// TIA Portal project "SemesterprosjektV7" (V20)

(* hardware
DEVICE "S7-1200 station_1"  S7-1200 Station
   slot 0: "Rack_0"  S7-1200 Rack  Rack  V1.0
   slot 1: "PLC_1"  CPU 1212C AC/DC/Rly  6ES7 212-1BD30-0XB0  V2.0
   slot 2: "AI 4x13BIT_1"  SM 1231 AI4  6ES7 231-4HD32-0XB0  V2.1
   slot 3: "AQ 2x14BIT_1"  SM 1232 AQ2  6ES7 232-4HB32-0XB0  V2.1
DEVICE "HMI_1"  KTP700 Basic PN
   slot 0: "HMI_1"  KTP700 Basic PN  6AV2 123-2GB03-0AX0  17.0.0.0
   slot 1: "HMI_RT_1"  KTP700 Basic PN  6AV2 123-2GB03-0AX0  17.0.0.0
   slot 5: "HMI_1.IE_CP_1"  PROFINET Interface  17.0.0.0
      slot 1: "PROFINET Interface_1"  PROFINET Interface
         slot 1: "Port_1"  Port
*)

// ===== PLC "PLC_1"  CPU 1212C AC/DC/Rly =====

VAR_GLOBAL   // PLC tag table "Default tag table"
   "AI2+" AT %IW100 : Int;
   "AQ1_PÅDRAG_PUMP1" AT %QW112 : Int;
   "AQ2" AT %QW114 : Int;
   "DI_EM_STOP" AT %I0.0 : Bool;
   "DQ_START_PUMP1" AT %Q0.0 : Bool;
   "DI_LS_Tørrkjøringsvern" AT %I0.1 : Bool;
   "DI_Reset_EM_STOP" AT %I0.2 : Bool;
   "DQ_Lys_EM_STOP" AT %Q0.1 : Bool;
END_VAR

// folder: Equipment

TYPE "UDT_Mal"
   STRUCT
      CFG : Struct   // Configuration Data
         Spare : Bool;
      END_STRUCT;
      Sts : Struct   // Status Data
         Spare : Bool;
      END_STRUCT;
      Cmd : Struct   // Command and request Data
         Spare : Bool;
      END_STRUCT;
      Par : Struct   // Parameter Data
         Spare : Bool;
      END_STRUCT;
      Fit : Struct   // Warning and alarm triggers
         Spare : Bool;
      END_STRUCT;
   END_STRUCT;
END_TYPE

TYPE "UDT_Pump_Control"
   STRUCT
      CFG : Struct   // Configuration Data
         Spare : Bool;
      END_STRUCT;
      Sts : Struct   // Status Data
         Spare : Bool;
      END_STRUCT;
      Cmd : Struct   // Command and request Data
         Start_Pump : Bool;
         Stop_Pump : Bool;
         EM_Stop : Bool;
      END_STRUCT;
      Par : Struct   // Parameter Data
         Pådrag_Inn : Real;
      END_STRUCT;
      Fit : Struct   // Warning and alarm triggers
         Feil : Bool;
      END_STRUCT;
   END_STRUCT;
END_TYPE

TYPE "UDT_Level_Transmitter"
   STRUCT
      CFG : Struct   // Configuration Data
         Spare : Bool;
      END_STRUCT;
      Sts : Struct   // Status Data
         Spare : Bool;
      END_STRUCT;
      Cmd : Struct   // Command and request Data
         Spare : Bool;
      END_STRUCT;
      Par : Struct   // Parameter Data
         EU_Value_Out : Real;
      END_STRUCT;
      Fit : Struct   // Warning and alarm triggers
         Feil : Bool;
         Spare : Bool;
      END_STRUCT;
   END_STRUCT;
END_TYPE

// folder: Machine

TYPE "UDT_HMI"
   STRUCT
      CFG : Struct   // Configuration Data
         Spare : Bool;
      END_STRUCT;
      Sts : Struct   // Status Data
         HMI_Level_PV : Real;
      END_STRUCT;
      Cmd : Struct   // Command and request Data
         HMI_Auto : Bool;
         HMI_Manuell : Bool;
         HMI_Start_Pump1 : Bool;
         HMI_Stop_Pump1 : Bool;
         HMI_Knapp_Auto : Bool;
         HMI_Knapp_Manuell : Bool;
         HMI_Knapp_Start_Pump1 : Bool;
         HMI_Knapp_Stop_Pump1 : Bool;
         Spare : Bool;
      END_STRUCT;
      Par : Struct   // Parameter Data
         HMI_P_Gain : Real;
         HMI_Ti : Real;
         HMI_Td : Real;
         HMI_Manual_Speed_Ref_P1 : Real;
         HMI_Level_SP : Real;
         HMI_EU_Min : Real;
         HMI_EU_Max : Real;
         HMI_Anti_Windup : Bool;
         Spare : Bool;
      END_STRUCT;
      Fit : Struct   // Warning and alarm triggers
         HMI_EM_Stop_Alarm : Bool;
         HMI_LS_Activated : Bool;
         HMI_Pump_Fault_Timer_SP : Time;
         HMI_Pump_Fault : Bool;
         Spare : Bool;
      END_STRUCT;
   END_STRUCT;
END_TYPE

// folder: (top level)

DATA_BLOCK "LT01"   // DB3
{ S7_Optimized_Access := 'TRUE' }
VERSION : 0.1
// stored: InstanceOfName Level_Transmitter
"Level_Transmitter"
BEGIN
END_DATA_BLOCK

DATA_BLOCK "Analog_Data"   // DB4
{ S7_Optimized_Access := 'TRUE' }
VERSION : 0.1
   VAR
      Raw_Value : Real;
      Output : Real;
      EU_Min : Real;
      EU_Max : Real;
   END_VAR
BEGIN
END_DATA_BLOCK

DATA_BLOCK "Pump1_Control_DB"   // DB6
{ S7_Optimized_Access := 'TRUE' }
VERSION : 0.1
// stored: InstanceOfName Pump_Control
"Pump_Control"
BEGIN
END_DATA_BLOCK

DATA_BLOCK "Machine01_DB"   // DB7
{ S7_Optimized_Access := 'TRUE' }
VERSION : 0.1
// stored: InstanceOfName Machine01
"Machine01"
BEGIN
END_DATA_BLOCK

DATA_BLOCK "Regulator_DB"   // DB9
{ S7_Optimized_Access := 'TRUE' }
VERSION : 0.1
// stored: InstanceOfName Regulator
"Regulator"
BEGIN
END_DATA_BLOCK

// folder: Global_Data

DATA_BLOCK "DB_Machine"   // DB1
{ S7_Optimized_Access := 'TRUE' }
VERSION : 0.1
   VAR
      HMI_Control : "UDT_HMI";
   END_VAR
BEGIN
END_DATA_BLOCK

DATA_BLOCK "DB_Equipment"   // DB2
{ S7_Optimized_Access := 'TRUE' }
VERSION : 0.1
   VAR
      Pump1_Control : "UDT_Pump_Control";
      LT01_Control : "UDT_Level_Transmitter";
      HMI_Control : "UDT_HMI";
   END_VAR
BEGIN
END_DATA_BLOCK

// folder: System blocks/Program resources

DATA_BLOCK "EM_Stop_TON_DB"   // DB5
{ S7_Optimized_Access := 'TRUE' }
AUTHOR : Simatic
FAMILY : IEC
NAME : IEC_TMR
VERSION : 1.0
// stored: InstanceOfName IEC_TIMER
"IEC_TIMER"
BEGIN
END_DATA_BLOCK

DATA_BLOCK "EM_Stop_TOF_DB"   // DB10
{ S7_Optimized_Access := 'TRUE' }
AUTHOR : Simatic
FAMILY : IEC
NAME : IEC_TMR
VERSION : 1.0
// stored: InstanceOfName IEC_TIMER
"IEC_TIMER"
BEGIN
END_DATA_BLOCK

DATA_BLOCK "Pump_Fault_Timer_DB"   // DB11
{ S7_Optimized_Access := 'TRUE' }
AUTHOR : Simatic
FAMILY : IEC
NAME : IEC_TMR
VERSION : 1.0
// stored: InstanceOfName IEC_TIMER
"IEC_TIMER"
BEGIN
END_DATA_BLOCK

// folder: (top level)

ORGANIZATION_BLOCK "Main"   // OB1, LAD, ProgramCycle
TITLE = "Main Program Sweep (Cycle)"
{ S7_Optimized_Access := 'TRUE' }
VERSION : 0.1
BEGIN
END_ORGANIZATION_BLOCK

ORGANIZATION_BLOCK "Machine"   // OB123, LAD, ProgramCycle
TITLE = "Main Program Sweep (Cycle)"
{ S7_Optimized_Access := 'TRUE' }
VERSION : 0.1
BEGIN

REGION Network 1
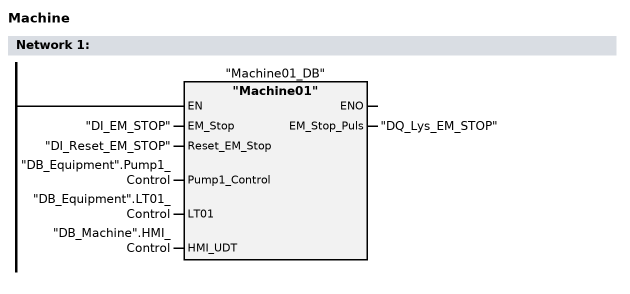
   RUNG wire#powerrail
      "Machine01_DB"(EM_Stop := "DI_EM_STOP", Reset_EM_Stop := "DI_Reset_EM_STOP", Pump1_Control := "DB_Equipment".Pump1_Control, LT01 := "DB_Equipment".LT01_Control, HMI_UDT := "DB_Machine".HMI_Control, EM_Stop_Puls => "DQ_Lys_EM_STOP")
   END_RUNG
   // the same network as SCL:
   "Machine01_DB"(EM_Stop := "DI_EM_STOP",   // "Machine01"
                  Reset_EM_Stop := "DI_Reset_EM_STOP",
                  Pump1_Control := "DB_Equipment".Pump1_Control,
                  LT01 := "DB_Equipment".LT01_Control,
                  HMI_UDT := "DB_Machine".HMI_Control,
                  EM_Stop_Puls => "DQ_Lys_EM_STOP");
END_REGION
END_ORGANIZATION_BLOCK

ORGANIZATION_BLOCK "Equipment"   // OB124, LAD, ProgramCycle
TITLE = "Main Program Sweep (Cycle)"
{ S7_Optimized_Access := 'TRUE' }
VERSION : 0.1
BEGIN

REGION Network 1
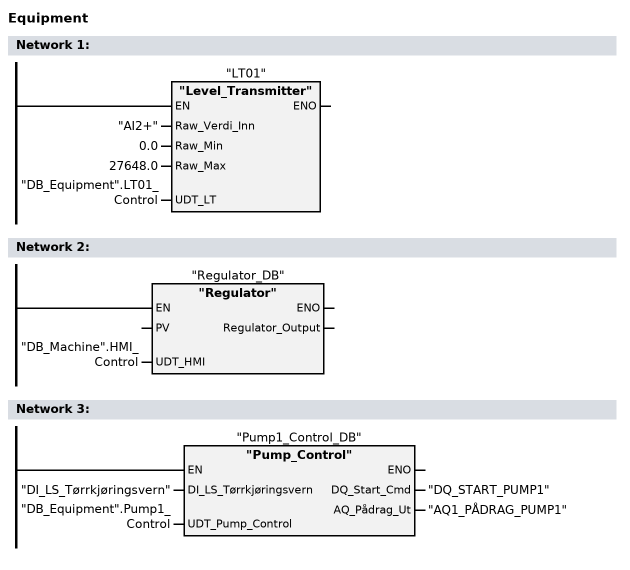
   RUNG wire#powerrail
      "LT01"(Raw_Verdi_Inn := "AI2+", Raw_Min := 0.0, Raw_Max := 27648.0, UDT_LT := "DB_Equipment".LT01_Control)
   END_RUNG
   // the same network as SCL:
   "LT01"(Raw_Verdi_Inn := "AI2+", Raw_Min := 0.0, Raw_Max := 27648.0, UDT_LT := "DB_Equipment".LT01_Control);   // "Level_Transmitter"
END_REGION

REGION Network 2
   RUNG wire#powerrail
      "Regulator_DB"(PV :=, UDT_HMI := "DB_Machine".HMI_Control, Regulator_Output =>)
   END_RUNG
   // the same network as SCL:
   "Regulator_DB"(UDT_HMI := "DB_Machine".HMI_Control);   // "Regulator"
END_REGION

REGION Network 3
   RUNG wire#powerrail
      "Pump1_Control_DB"(DI_LS_Tørrkjøringsvern := "DI_LS_Tørrkjøringsvern", UDT_Pump_Control := "DB_Equipment".Pump1_Control, DQ_Start_Cmd => "DQ_START_PUMP1", AQ_Pådrag_Ut => "AQ1_PÅDRAG_PUMP1")
   END_RUNG
   // the same network as SCL:
   "Pump1_Control_DB"(DI_LS_Tørrkjøringsvern := "DI_LS_Tørrkjøringsvern",   // "Pump_Control"
                      UDT_Pump_Control := "DB_Equipment".Pump1_Control,
                      DQ_Start_Cmd => "DQ_START_PUMP1",
                      AQ_Pådrag_Ut => "AQ1_PÅDRAG_PUMP1");
END_REGION
END_ORGANIZATION_BLOCK

// folder: Equipment

FUNCTION_BLOCK "Pump_Control"   // FB2, LAD
{ S7_Optimized_Access := 'TRUE' }
VERSION : 0.1
   VAR_INPUT
      DI_LS_Tørrkjøringsvern : Bool;
   END_VAR
   VAR_OUTPUT
      DQ_Start_Cmd : Bool;
      AQ_Pådrag_Ut : Int;
   END_VAR
   VAR_IN_OUT
      UDT_Pump_Control : "UDT_Pump_Control";
   END_VAR
   VAR
      Tmp_Start_Cmd : Bool;
      Tmp_Pådrag_Ut_Real : Real;
      Temp_Verdi : Real;
      Tmp_Pådrag_Ut_Int : Real;
   END_VAR
BEGIN

REGION Network 1
   // Start Pumpe og stopp kriterier
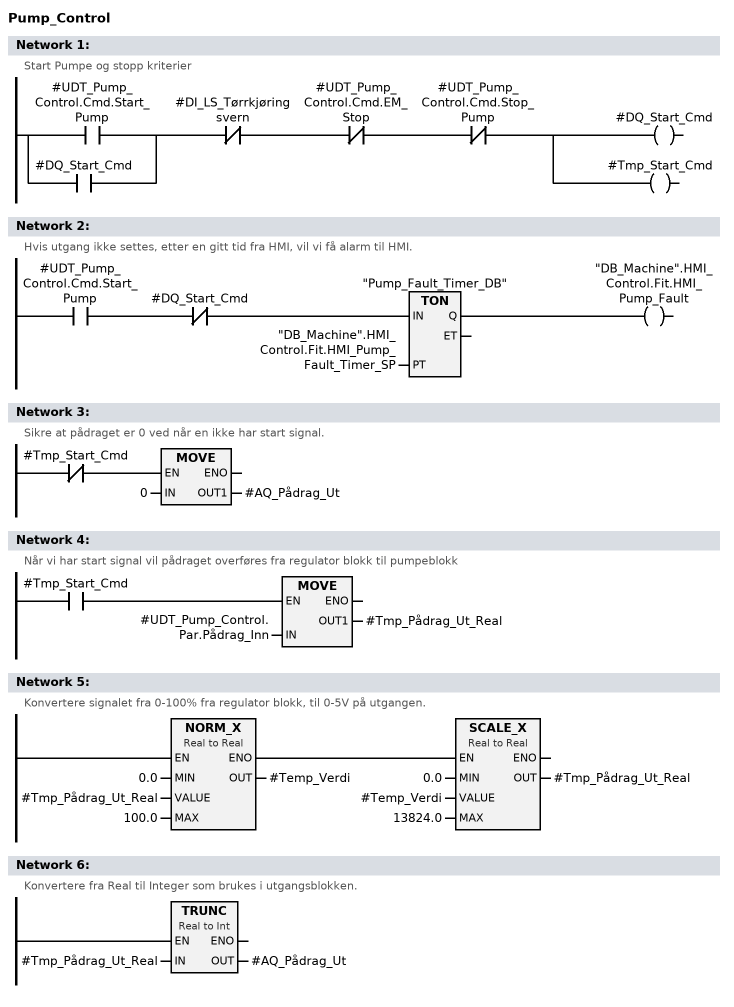
   RUNG wire#powerrail
      Contact( #UDT_Pump_Control.Cmd.Start_Pump )
      wire#w1
      I_Contact( #DI_LS_Tørrkjøringsvern )
      I_Contact( #UDT_Pump_Control.Cmd.EM_Stop )
      I_Contact( #UDT_Pump_Control.Cmd.Stop_Pump )
      wire#w2
      Coil( #DQ_Start_Cmd )
   END_RUNG
   RUNG wire#powerrail
      Contact( #DQ_Start_Cmd )
   END_RUNG wire#w1
   RUNG wire#w2
      Coil( #Tmp_Start_Cmd )
   END_RUNG
   // the same network as SCL:
   #DQ_Start_Cmd := (#UDT_Pump_Control.Cmd.Start_Pump OR #DQ_Start_Cmd) AND NOT #DI_LS_Tørrkjøringsvern AND NOT #UDT_Pump_Control.Cmd.EM_Stop AND NOT #UDT_Pump_Control.Cmd.Stop_Pump;
   #Tmp_Start_Cmd := #DQ_Start_Cmd;
END_REGION

REGION Network 2
   // Hvis utgang ikke settes, etter en gitt tid fra HMI, vil vi få alarm til HMI.
   "Pump_Fault_Timer_DB".TON(IN := #UDT_Pump_Control.Cmd.Start_Pump AND NOT #DQ_Start_Cmd,
                           PT := "DB_Machine".HMI_Control.Fit.HMI_Pump_Fault_Timer_SP);
   "DB_Machine".HMI_Control.Fit.HMI_Pump_Fault := "Pump_Fault_Timer_DB".Q;
END_REGION

REGION Network 3
   // Sikre at pådraget er 0 ved når en ikke har start signal.
   RUNG wire#powerrail
      I_Contact( #Tmp_Start_Cmd )
      { S7_GenerateENO := "TRUE" } Move(in := 0, out1 => #AQ_Pådrag_Ut)
   END_RUNG
   // the same network as SCL:
   IF NOT #Tmp_Start_Cmd THEN #AQ_Pådrag_Ut := 0; END_IF;
END_REGION

REGION Network 4
   // Når vi har start signal vil pådraget overføres fra regulator blokk til pumpeblokk
   RUNG wire#powerrail
      Contact( #Tmp_Start_Cmd )
      { S7_GenerateENO := "TRUE" } Move(in := #UDT_Pump_Control.Par.Pådrag_Inn, out1 => #Tmp_Pådrag_Ut_Real)
   END_RUNG
   // the same network as SCL:
   IF #Tmp_Start_Cmd THEN #Tmp_Pådrag_Ut_Real := #UDT_Pump_Control.Par.Pådrag_Inn; END_IF;
END_REGION

REGION Network 5
   // Konvertere signalet fra 0-100% fra regulator blokk, til 0-5V på utgangen.
   RUNG wire#powerrail
      { S7_Templates := "[SrcType := Real, DestType := Real]"; S7_GenerateENO := "TRUE" } Normalize(min := 0.0, value := #Tmp_Pådrag_Ut_Real, max := 100.0, out => #Temp_Verdi)
      { S7_Templates := "[SrcType := Real, DestType := Real]"; S7_GenerateENO := "TRUE" } Scale(min := 0.0, value := #Temp_Verdi, max := 13824.0, out => #Tmp_Pådrag_Ut_Real)
   END_RUNG
   // the same network as SCL:
   // ENO of a box is taken as its EN; it also drops when the box reports an error
   #Temp_Verdi := NORM_X(MIN := 0.0, VALUE := #Tmp_Pådrag_Ut_Real, MAX := 100.0);
   #Tmp_Pådrag_Ut_Real := SCALE_X(MIN := 0.0, VALUE := #Temp_Verdi, MAX := 13824.0);
END_REGION

REGION Network 6
   // Konvertere fra Real til Integer som brukes i utgangsblokken.
   RUNG wire#powerrail
      { S7_Templates := "[SrcType := Real, DestType := Int]"; S7_GenerateENO := "TRUE" } Trunc(in := #Tmp_Pådrag_Ut_Real, out => #AQ_Pådrag_Ut)
   END_RUNG
   // the same network as SCL:
   #AQ_Pådrag_Ut := TRUNC(#Tmp_Pådrag_Ut_Real);
END_REGION
END_FUNCTION_BLOCK

FUNCTION_BLOCK "Level_Transmitter"   // FB3, LAD
{ S7_Optimized_Access := 'TRUE' }
VERSION : 0.1
   VAR_INPUT
      Raw_Verdi_Inn : Int;
      Raw_Min : Real;
      Raw_Max : Real;
   END_VAR
   VAR_IN_OUT
      UDT_LT : "UDT_Level_Transmitter";
   END_VAR
   VAR_TEMP
      Convert_Value : Real;
      Raw_Value_Real : Real;
   END_VAR
BEGIN

REGION Network 1
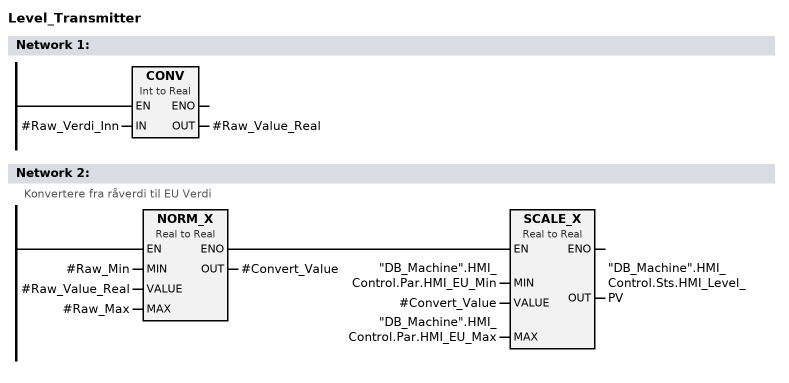
   RUNG wire#powerrail
      { S7_Templates := "[SrcType := Int, DestType := Real]"; S7_GenerateENO := "TRUE" } Convert(in := #Raw_Verdi_Inn, out => #Raw_Value_Real)
   END_RUNG
   // the same network as SCL:
   #Raw_Value_Real := INT_TO_REAL(#Raw_Verdi_Inn);
END_REGION

REGION Network 2
   // Konvertere fra råverdi til EU Verdi
   RUNG wire#powerrail
      { S7_Templates := "[SrcType := Real, DestType := Real]"; S7_GenerateENO := "TRUE" } Normalize(min := #Raw_Min, value := #Raw_Value_Real, max := #Raw_Max, out => #Convert_Value)
      { S7_Templates := "[SrcType := Real, DestType := Real]"; S7_GenerateENO := "TRUE" } Scale(min := "DB_Machine".HMI_Control.Par.HMI_EU_Min, value := #Convert_Value, max := "DB_Machine".HMI_Control.Par.HMI_EU_Max, out => "DB_Machine".HMI_Control.Sts.HMI_Level_PV)
   END_RUNG
   // the same network as SCL:
   // ENO of a box is taken as its EN; it also drops when the box reports an error
   #Convert_Value := NORM_X(MIN := #Raw_Min, VALUE := #Raw_Value_Real, MAX := #Raw_Max);
   "DB_Machine".HMI_Control.Sts.HMI_Level_PV := SCALE_X(MIN := "DB_Machine".HMI_Control.Par.HMI_EU_Min, VALUE := #Convert_Value, MAX := "DB_Machine".HMI_Control.Par.HMI_EU_Max);
END_REGION
END_FUNCTION_BLOCK

FUNCTION_BLOCK "ØL_PID"   // FB4, LAD
{ S7_Optimized_Access := 'TRUE' }
VERSION : 0.1
   VAR_INPUT
      SP : LReal;   // // NRM / SIU Setpoint
      PV : LReal;   // // NRM / SIU Process Value
      Bias : LReal;   // // NRM Bias Value
      I_SP : LReal;   // // NRM Setpoint for integrator value
      I_SP_Cmd : Bool;   // // TRUE: Load I_SP
      Suspend : Bool;   // // TRUE: Suspends operation
   END_VAR
   VAR_OUTPUT
      EV : LReal;   // // NRM / SIU Error Value
      CV : LReal;   // // NRM Control Value
   END_VAR
BEGIN
END_FUNCTION_BLOCK

FUNCTION_BLOCK "Regulator"   // FB5, LAD
{ S7_Optimized_Access := 'TRUE' }
VERSION : 0.1
   VAR_INPUT
      PV : Real;
   END_VAR
   VAR_OUTPUT
      Regulator_Output : Real;
   END_VAR
   VAR_IN_OUT
      UDT_HMI : "UDT_HMI";
   END_VAR
   VAR
      Convert_Value : Real;
      "Regulator_PV_%" : Real;
   END_VAR
BEGIN

REGION Network 2
   // Konvertere fra råverdi til EU Verdi
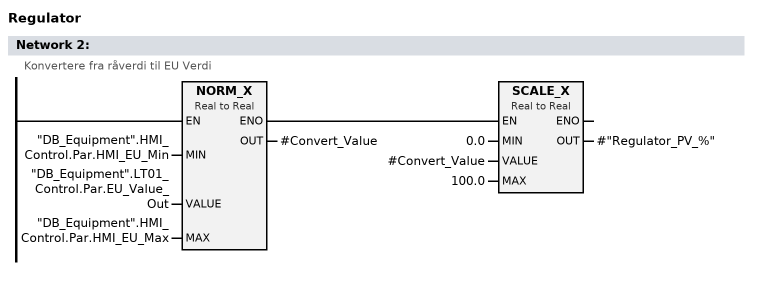
   RUNG wire#powerrail
      { S7_Templates := "[SrcType := Real, DestType := Real]"; S7_GenerateENO := "TRUE" } Normalize(min := "DB_Equipment".HMI_Control.Par.HMI_EU_Min, value := "DB_Equipment".LT01_Control.Par.EU_Value_Out, max := "DB_Equipment".HMI_Control.Par.HMI_EU_Max, out => #Convert_Value)
      { S7_Templates := "[SrcType := Real, DestType := Real]"; S7_GenerateENO := "TRUE" } Scale(min := 0.0, value := #Convert_Value, max := 100.0, out => #"Regulator_PV_%")
   END_RUNG
   // the same network as SCL:
   // ENO of a box is taken as its EN; it also drops when the box reports an error
   #Convert_Value := NORM_X(MIN := "DB_Equipment".HMI_Control.Par.HMI_EU_Min, VALUE := "DB_Equipment".LT01_Control.Par.EU_Value_Out, MAX := "DB_Equipment".HMI_Control.Par.HMI_EU_Max);
   #"Regulator_PV_%" := SCALE_X(MIN := 0.0, VALUE := #Convert_Value, MAX := 100.0);
END_REGION
END_FUNCTION_BLOCK

// folder: Machine

FUNCTION_BLOCK "Machine01"   // FB1, LAD
{ S7_Optimized_Access := 'TRUE' }
VERSION : 0.1
   VAR_INPUT
      EM_Stop : Bool;
      Reset_EM_Stop : Bool;
   END_VAR
   VAR_OUTPUT
      EM_Stop_Puls : Bool;
   END_VAR
   VAR_IN_OUT
      Pump1_Control : "UDT_Pump_Control";
      LT01 : "UDT_Level_Transmitter";
      HMI_UDT : "UDT_HMI";
   END_VAR
   VAR
      Tmp_EM_Stop : Bool;
      Tmp_Enable_PID : Bool;
      Tmp_Blink_Off : Bool;
      Tmp_Blink_On : Bool;
   END_VAR
BEGIN

REGION Network 1
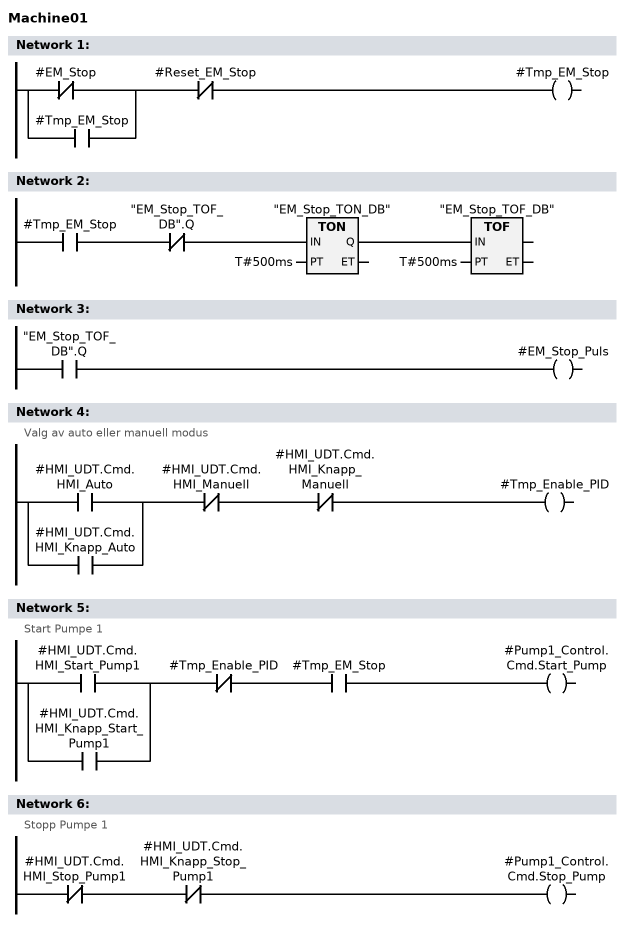
   RUNG wire#powerrail
      I_Contact( #EM_Stop )
      wire#w1
      I_Contact( #Reset_EM_Stop )
      Coil( #Tmp_EM_Stop )
   END_RUNG
   RUNG wire#powerrail
      Contact( #Tmp_EM_Stop )
   END_RUNG wire#w1
   // the same network as SCL:
   #Tmp_EM_Stop := (NOT #EM_Stop OR #Tmp_EM_Stop) AND NOT #Reset_EM_Stop;
END_REGION

REGION Network 2
   "EM_Stop_TON_DB".TON(IN := #Tmp_EM_Stop AND NOT "EM_Stop_TOF_DB".Q, PT := T#500ms);
   "EM_Stop_TOF_DB".TOF(IN := "EM_Stop_TON_DB".Q, PT := T#500ms);
END_REGION

REGION Network 3
   RUNG wire#powerrail
      Contact( "EM_Stop_TOF_DB".Q )
      Coil( #EM_Stop_Puls )
   END_RUNG
   // the same network as SCL:
   #EM_Stop_Puls := "EM_Stop_TOF_DB".Q;
END_REGION

REGION Network 4
   // Valg av auto eller manuell modus
   RUNG wire#powerrail
      Contact( #HMI_UDT.Cmd.HMI_Auto )
      wire#w1
      I_Contact( #HMI_UDT.Cmd.HMI_Manuell )
      I_Contact( #HMI_UDT.Cmd.HMI_Knapp_Manuell )
      Coil( #Tmp_Enable_PID )
   END_RUNG
   RUNG wire#powerrail
      Contact( #HMI_UDT.Cmd.HMI_Knapp_Auto )
   END_RUNG wire#w1
   // the same network as SCL:
   #Tmp_Enable_PID := (#HMI_UDT.Cmd.HMI_Auto OR #HMI_UDT.Cmd.HMI_Knapp_Auto) AND NOT #HMI_UDT.Cmd.HMI_Manuell AND NOT #HMI_UDT.Cmd.HMI_Knapp_Manuell;
END_REGION

REGION Network 5
   // Start Pumpe 1
   RUNG wire#powerrail
      Contact( #HMI_UDT.Cmd.HMI_Start_Pump1 )
      wire#w1
      I_Contact( #Tmp_Enable_PID )
      Contact( #Tmp_EM_Stop )
      Coil( #Pump1_Control.Cmd.Start_Pump )
   END_RUNG
   RUNG wire#powerrail
      Contact( #HMI_UDT.Cmd.HMI_Knapp_Start_Pump1 )
   END_RUNG wire#w1
   // the same network as SCL:
   #Pump1_Control.Cmd.Start_Pump := (#HMI_UDT.Cmd.HMI_Start_Pump1 OR #HMI_UDT.Cmd.HMI_Knapp_Start_Pump1) AND NOT #Tmp_Enable_PID AND #Tmp_EM_Stop;
END_REGION

REGION Network 6
   // Stopp Pumpe 1
   RUNG wire#powerrail
      I_Contact( #HMI_UDT.Cmd.HMI_Stop_Pump1 )
      I_Contact( #HMI_UDT.Cmd.HMI_Knapp_Stop_Pump1 )
      Coil( #Pump1_Control.Cmd.Stop_Pump )
   END_RUNG
   // the same network as SCL:
   #Pump1_Control.Cmd.Stop_Pump := NOT #HMI_UDT.Cmd.HMI_Stop_Pump1 AND NOT #HMI_UDT.Cmd.HMI_Knapp_Stop_Pump1;
END_REGION
END_FUNCTION_BLOCK

(* ===== HMI "HMI_RT_1" =====
system functions are stored by id; their names below are inferred from use
connection "HMI_Connection_1": ETHERNET, SMART_S7_1200_OMS

HMI tags "HMI_Tags"
   "Knapp_HMI_Stop_Pump1" : Bool = PLC DB_Machine.HMI_Control.Cmd.HMI_Knapp_Stop_Pump1 AT %DB1.DBX0.0, 1 s
   "HMI_Manuell" : Bool = PLC DB_Machine.HMI_Control.Cmd.HMI_Manuell AT %DB1.DBX0.0, 1 s
   "HMI_Start_Pump1" : Bool = PLC DB_Machine.HMI_Control.Cmd.HMI_Start_Pump1 AT %DB1.DBX0.0, 1 s
   "Knapp_HMI_Auto" : Bool = PLC DB_Machine.HMI_Control.Cmd.HMI_Knapp_Auto AT %DB1.DBX0.0, 1 s
   "HMI_Auto" : Bool = PLC DB_Machine.HMI_Control.Cmd.HMI_Auto AT %DB1.DBX0.0, 1 s
   "Knapp_HMI_Manuell" : Bool = PLC DB_Machine.HMI_Control.Cmd.HMI_Knapp_Manuell AT %DB1.DBX0.0, 1 s
   "Knapp_HMI_Start_Pump1" : Bool = PLC DB_Machine.HMI_Control.Cmd.HMI_Knapp_Start_Pump1 AT %DB1.DBX0.0, 1 s
   "Tag_ScreenNumber_1" : UInt, internal
   "HMI_Stop_Pump1" : Bool = PLC DB_Machine.HMI_Control.Cmd.HMI_Stop_Pump1 AT %DB1.DBX0.0, 1 s
   "PID_Compact_1_Output" : Real = PLC PID_Compact_1.Output, 1 s
   "PID_Compact_1_Setpoint" : Real = PLC PID_Compact_1.Setpoint, 1 s

Template "Template_1" 800x480
   Button "Exit" at 714,429 size 71x50; TextOff 'Exit'; PictureOff "ExitRuntime_KTP700_Basic_PN_TR"; PictureOn "ExitRuntime_KTP700_Basic_PN_TR"
      on Release: StopRuntime(0)
   Button "Log on" at 614,429 size 71x50; TextOff 'Log on'; PictureOff "Login_KTP700_Basic_PN_TR"; PictureOn "Login_KTP700_Basic_PN_TR"
      on Release: function_a2a04561()
   Button "Template_Button" at 514,429 size 71x50; TextOff 'Text'
   Button "Template_Button_1" at 414,429 size 71x50; TextOff 'Text'
   Button "Template_Button_2" at 314,429 size 71x50; TextOff 'Text'
   Button "Template_Button_3" at 214,429 size 71x50; TextOff 'Text'
   Button "Alarms" at 114,429 size 71x50; TextOff 'Alarms'; PictureOff "AlarmDisplay_KTP700_Basic_PN_TR"; PictureOn "AlarmDisplay_KTP700_Basic_PN_TR"
      on Release: function_ef3f5d25("Alarm window_Unacknowledged", -1)
   Button "Start screen" at 14,429 size 71x50; TextOff 'Start screen'; PictureOff "NavigateHome_KTP700_Basic_PN_TR"; PictureOn "NavigateHome_KTP700_Basic_PN_TR"
      on Release: ActivateScreen("Root screen", 0)
   DateTimeField "HmiScreenItemData" at 695,25 size 105x25
   DateTimeField "HmiScreenItemData_1" at 695,0 size 105x25
   GraphicView "Logo" at 0,0 size 91x51; Picture "Logo of HMI_1"

screen "Root screen" 800x480, template "Template_1"
   on GenerateScreen: SetTag("HMI_Manuell", 1)
   TextField "HmiScreenItemData_3" at 107,58 size 640x25; Text 'Welcome to HMI_1 (KTP700 Basic+ PN)!'
   Button "HmiScreenItemData" at 36,87 size 159x47; TextOff 'Screen0'; PictureOff "Navigates to Screen0 for KTP700 Basic+ PN 17.0.0.0"; PictureOn "Navigates to Screen0 for KTP700 Basic+ PN 17.0.0.0"
      on Release: ActivateScreen("Screen0", 0)
   Button "HmiScreenItemData_1" at 36,146 size 159x47; TextOff 'Screen2'; PictureOff "Navigates to Screen2 for KTP700 Basic+ PN 17.0.0.0"; PictureOn "Navigates to Screen2 for KTP700 Basic+ PN 17.0.0.0"
      on Release: ActivateScreen("Screen2", 0)
   Button "HmiScreenItemData_2" at 36,205 size 159x47; TextOff 'Screen3'; PictureOff "Navigates to Screen3 for KTP700 Basic+ PN 17.0.0.0"; PictureOn "Navigates to Screen3 for KTP700 Basic+ PN 17.0.0.0"
      on Release: ActivateScreen("Screen3", 0)
   Button "HmiScreenItemData_4" at 36,264 size 159x47; TextOff 'System screens'; PictureOff "Navigates to System screens for KTP700 Basic+ PN 17.0.0.0"; PictureOn "Navigates to System screens for KTP700 Basic+ PN 17.0.0.0"
      on Release: ActivateScreen("System screens", 0)
   Button "Button_1" at 233,99 size 104x35; TextOff 'AUTO'
      on Click: ResetBit("HMI_Manuell"); SetBit("HMI_Auto")
   Button "Button_2" at 233,158 size 104x35; TextOff 'MANUELL'
      on Click: ResetBit("HMI_Auto"); SetBit("HMI_Manuell")
   Button "Button_3" at 389,99 size 164x35; TextOff 'START PUMP 1'
      on Click: ResetBit("HMI_Stop_Pump1"); SetBit("HMI_Start_Pump1")
   Button "Button_4" at 389,158 size 164x35; TextOff 'STOP PUMP 1'
      on Click: ResetBit("HMI_Start_Pump1"); SetBit("HMI_Stop_Pump1")
   IOField "I/O field_1" at 471,272 size 82x39; FormatPattern s999999999.999
      ProcessValue <- "PID_Compact_1_Output"
   IOField "I/O field_2" at 233,272 size 82x39; FormatPattern s999999999.999
      ProcessValue <- "PID_Compact_1_Setpoint"

screen "Screen0" 800x480, template "Template_1"
   on GenerateScreen: SetTag("Knapp_HMI_Stop_Pump1", 2)
   TextField "HmiScreenItemData" at 80,225 size 640x25; Text 'Screen0'
   Button "Back" at 1,52 size 159x47; TextOff 'Back'
      on Release: ActivateScreen("Root screen", 0)

screen "Screen2" 800x480, template "Template_1"
   on GenerateScreen: SetTag("Knapp_HMI_Stop_Pump1", 3)
   TextField "HmiScreenItemData" at 80,225 size 640x25; Text 'Screen2'
   Button "Back" at 1,52 size 159x47; TextOff 'Back'
      on Release: ActivateScreen("Root screen", 0)

screen "Screen3" 800x480, template "Template_1"
   on GenerateScreen: SetTag("Knapp_HMI_Stop_Pump1", 4)
   TextField "HmiScreenItemData" at 80,225 size 640x25; Text 'Screen3'
   Button "Back" at 1,52 size 159x47; TextOff 'Back'
      on Release: ActivateScreen("Root screen", 0)

screen "System screens" 800x480, template "Template_1"
   on GenerateScreen: SetTag("Knapp_HMI_Stop_Pump1", 5)
   Button "Back" at 1,52 size 159x47; TextOff 'Back'
      on Release: ActivateScreen("Root screen", 0)
   Button "HmiScreenItemData" at 36,146 size 159x47; TextOff 'SIMATIC PLC system diagnos...'; PictureOff "Navigates to SIMATIC PLC system diagnostics for KTP700 Basic+ PN 17.0.0.0"; PictureOn "Navigates to SIMATIC PLC system diagnostics for KTP700 Basic+ PN 17.0.0.0"
      on Release: ActivateScreen("SIMATIC PLC system diagnostics", 0)
   Button "HmiScreenItemData_1" at 36,205 size 159x47; TextOff 'Project information'; PictureOff "Navigates to Project information for KTP700 Basic+ PN 17.0.0.0"; PictureOn "Navigates to Project information for KTP700 Basic+ PN 17.0.0.0"
      on Release: ActivateScreen("Project information", 0)
   Button "HmiScreenItemData_2" at 36,264 size 159x47; TextOff 'User administration'; PictureOff "Navigates to User administration for KTP700 Basic+ PN 17.0.0.0"; PictureOn "Navigates to User administration for KTP700 Basic+ PN 17.0.0.0"
      on Release: ActivateScreen("User administration", 0)
   Button "HmiScreenItemData_3" at 36,323 size 159x47; TextOff 'System information'; PictureOff "Navigates to System information for KTP700 Basic+ PN 17.0.0.0"; PictureOn "Navigates to System information for KTP700 Basic+ PN 17.0.0.0"
      on Release: ActivateScreen("System information", 0)
   Button "HmiScreenItemData_4" at 207,146 size 159x47; TextOff 'Different jobs'; PictureOff "Navigates to Different jobs for KTP700 Basic+ PN 17.0.0.0"; PictureOn "Navigates to Different jobs for KTP700 Basic+ PN 17.0.0.0"
      on Release: ActivateScreen("Different jobs", 0)

screen "SIMATIC PLC system diagnostics" 800x480, template "Template_1"
   on GenerateScreen: SetTag("Knapp_HMI_Stop_Pump1", 6)
   SysDiagControl "HmiScreenItemData" at 1,100 size 796x321
   Button "Back" at 1,52 size 159x47; TextOff 'Back'
      on Release: ActivateScreen("System screens", 0)

screen "Project information" 800x480, template "Template_1"
   on GenerateScreen: SetTag("Knapp_HMI_Stop_Pump1", 7)
   TextField "HmiScreenItemData" at 35,102 size 171x28; Text 'Project name:'
   TextField "HmiScreenItemData_1" at 241,102 size 524x28; Text 'SemesterprosjektV2'
   TextField "HmiScreenItemData_2" at 35,132 size 171x28; Text 'Created on:'
   TextField "HmiScreenItemData_3" at 241,132 size 524x28; Text '11/7/2025 1:47:45 PM'
   TextField "HmiScreenItemData_4" at 35,162 size 171x28; Text 'Author:'
   TextField "HmiScreenItemData_5" at 241,162 size 524x28; Text 'Olav Eide'
   TextField "HmiScreenItemData_6" at 35,192 size 171x28; Text 'Description:'
   TextField "HmiScreenItemData_7" at 241,192 size 524x28; Text '(not configured)'
   Button "Back" at 1,52 size 159x47; TextOff 'Back'
      on Release: ActivateScreen("System screens", 0)

screen "User administration" 800x480, template "Template_1"
   on GenerateScreen: SetTag("Knapp_HMI_Stop_Pump1", 8)
   UserView "HmiScreenItemData" at 1,100 size 796x321
   Button "Back" at 1,52 size 159x47; TextOff 'Back'
      on Release: ActivateScreen("System screens", 0)

screen "System information" 800x480, template "Template_1"
   on GenerateScreen: SetTag("Knapp_HMI_Stop_Pump1", 9)
   TextField "HmiScreenItemData" at 35,102 size 171x28; Text 'HMI device type:'
   TextField "HmiScreenItemData_1" at 241,102 size 524x28; Text 'KTP700 Basic+ PN 17.0.0.0'
   TextField "HmiScreenItemData_2" at 35,132 size 171x28; Text 'Connection:'
   TextField "HmiScreenItemData_3" at 241,132 size 524x28; Text 'PROFINET (X1)'
   TextField "HmiScreenItemData_4" at 35,162 size 171x28; Text 'PLC:'
   TextField "HmiScreenItemData_5" at 241,162 size 524x28; Text 'SIMATIC S7 1200'
   Button "Back" at 1,52 size 159x47; TextOff 'Back'
      on Release: ActivateScreen("System screens", 0)

screen "Different jobs" 800x480, template "Template_1"
   on GenerateScreen: SetTag("Knapp_HMI_Stop_Pump1", 10)
   Button "Online" at 36,146 size 159x47; TextOff 'Online'
      on Release: function_bb44b551(0)
   Button "Offline" at 36,205 size 159x47; TextOff 'Offline'
      on Release: function_bb44b551(1)
   Button "Transfer" at 36,264 size 159x47; TextOff 'Transfer'
      on Release: function_bb44b551(2)
   Button "Toggle language" at 36,323 size 159x47; TextOff 'Toggle language'
      on Release: function_fb9197e8(-1)
   Button "Stop Runtime" at 207,146 size 159x47; TextOff 'Stop Runtime'
      on Release: StopRuntime(0)
   Button "Back" at 1,52 size 159x47; TextOff 'Back'
      on Release: ActivateScreen("System screens", 0)
*)